// TIA Portal project "THELMA3_200224" (V15.1)

(* hardware
DEVICE "S71500/ET200MP station_1"  S7-1500 station
   slot 0: "Rail_0"  Rack  6ES7 590-1***0-0AA0
   slot 0: "PM 190W 120/230VAC"  PM 190W 120/230VAC  6EP1333-4BA00
   slot 1: "THELMA3"  CPU 1515-2 PN  6ES7 515-2AM01-0AB0  V2.6
      slot 3: "CPU display_1"  6ES7591-1BA00-0AA0
   slot 2: "DI 16x24VDC HF_1"  DI 16x24VDC HF  6ES7 521-1BH00-0AB0  V2.2
   slot 3: "DQ 16x24VDC/0.5A HF_1"  DQ 16x24VDC/0.5A HF  6ES7 522-1BH01-0AB0  V1.1
   slot 4: "DQ 16x24VDC/0.5A HF_2"  DQ 16x24VDC/0.5A HF  6ES7 522-1BH01-0AB0  V1.1
DEVICE "GSD device_1"  GSD.Device.PN
   slot 0: "Rack"  Rack  V1.0
   slot 0: "ucm8-bag-thelma3"  DataMan 260  DMR-260#-#0  5.5.0
      slot 0: "DataMan 260"  DataMan 260
      slot 1: "Interface"  Interface
         slot 1: "Port 1"  Port 1
   slot 1: "Acquisition Control_1"  Acquisition Control
      slot 0: "Acquisition Control"  Acquisition Control
   slot 2: "Acquisition Status_1"  Acquisition Status
      slot 0: "Acquisition Status"  Acquisition Status
   slot 3: "Results Control_1"  Results Control
      slot 0: "Results Control"  Results Control
   slot 4: "Results Status_1"  Results Status
      slot 0: "Results Status"  Results Status
   slot 5: "Soft Event Control_1"  Soft Event Control
      slot 0: "Soft Event Control"  Soft Event Control
   slot 6: "User Data - 64 bytes_1"  User Data - 64 bytes
      slot 0: "User Data - 64 bytes"  User Data - 64 bytes
   slot 7: "Result Data - 64 bytes_1"  Result Data - 64 bytes
      slot 0: "Result Data - 64 bytes"  Result Data - 64 bytes
DEVICE "GSD device_2"  GSD.Device.PN
   slot 0: "Rack"  Rack  V1.0
   slot 0: "ucm8-box-thelma3"  DataMan 260  DMR-260#-#0  5.5.0
      slot 0: "DataMan 260"  DataMan 260
      slot 1: "Interface"  Interface
         slot 1: "Port 1"  Port 1
   slot 1: "Acquisition Control_1"  Acquisition Control
      slot 0: "Acquisition Control"  Acquisition Control
   slot 2: "Acquisition Status_1"  Acquisition Status
      slot 0: "Acquisition Status"  Acquisition Status
   slot 3: "Results Control_1"  Results Control
      slot 0: "Results Control"  Results Control
   slot 4: "Results Status_1"  Results Status
      slot 0: "Results Status"  Results Status
   slot 5: "Soft Event Control_1"  Soft Event Control
      slot 0: "Soft Event Control"  Soft Event Control
   slot 6: "User Data - 128 bytes_1"  User Data - 128 bytes
      slot 0: "User Data - 128 bytes"  User Data - 128 bytes
   slot 7: "Result Data - 128 bytes_1"  Result Data - 128 bytes
      slot 0: "Result Data - 128 bytes"  Result Data - 128 bytes
DEVICE "HMI_THELMA3"  TP700 Comfort
   slot 0: "HMI_THELMA3"  TP700 Comfort  6AV2 124-0GC01-0AX0  15.1.0.0
   slot 1: "HMI_RT_2"  TP700 Comfort  6AV2 124-0GC01-0AX0  15.1.0.0
   slot 5: "HMI_THELMA3.1"  PROFINET Interface  15.0.1.0
      slot 1: "PROFINET Interface_1"  PROFINET Interface
         slot 1: "Port_1"  Port
         slot 2: "Port_2"  Port
   slot 7: "HMI_THELMA3._CP_1"  MPI/DP Interface  15.0.1.0
*)

// ===== PLC "THELMA3"  CPU 1515-2 PN =====

VAR_GLOBAL   // PLC tag table "Default tag table"
   "TrigerSensor" AT %I10.7 : Bool;
   "x_BypassPlainCheck" AT %M500.0 : Bool;
   "x_Arikel1" AT %M500.1 : Bool;
   "x_Artikel2" AT %M500.2 : Bool;
   "x_Artikel3" AT %M500.3 : Bool;
   "x_Artikel4" AT %M500.4 : Bool;
   "x_Simulacia_NoveData" AT %M505.0 : Bool;
   "x_Simulacia_Error" AT %M505.6 : Bool;
   "Kamera_odpojena" AT %M18.0 : Bool;
   "ArticleChangingBag" AT %M10.0 : Bool;
   "ArticleChangingBox" AT %M10.1 : Bool;
   "Reader2_Trigger_DelayTime" AT %MD68 : Time;
   "CON_HF_CommandTrigBatch" AT %M120.0 : Bool;
   "CON_HF_CommandTrig" AT %M120.1 : Bool;
   "CON_HF_CommandTrigBatchCon" AT %M120.2 : Bool;
   "CON_HF_CommandTrigAgainBatch" AT %M120.6 : Bool;
   "CON_HF_CommandTrigAgain" AT %M120.7 : Bool;
   "FirstScan" AT %M1.0 : Bool;
   "DiagStatusUpdate" AT %M1.1 : Bool;
   "TimeSynchPeriod" AT %MD64 : Time;
   "AlarmCheckPeriod" AT %MD60 : Time;
   "FaultByte1" AT %MB100 : Byte;
   "FaultByte2" AT %MB101 : Byte;
   "DelayTimeReader" AT %MD13 : Time;
   "CON_PrinterSelection" AT %M8.0 : Bool;
   "TRP_ErrorIP" AT %M105.0 : Bool;
   "TRP_CommError" AT %M105.1 : Bool;
   "TRP_HF_CommandTrig" AT %M121.1 : Bool;
   "TRP_ConnectHMI" AT %M121.4 : Bool;
   "TRP_HF_CommandTrigAgain" AT %M121.7 : Bool;
   "TRP_Inverse" AT %M140.0 : Bool;
   "TRP_Label" AT %M140.1 : Bool;
   "FaultByte3" AT %MB102 : Byte;
   "ResetFaults(1)" AT %M8.1 : Bool;
   "ResetCounters" AT %M8.2 : Bool;
   "CON_PrinterConnection" AT %M8.3 : Bool;
   "CON_ConnectHMI" AT %M120.4 : Bool;
   "System_Byte" AT %MB1 : Byte;
   "AlwaysTRUE" AT %M1.2 : Bool;
   "AlwaysFALSE" AT %M1.3 : Bool;
   "ResetResultAck" AT %M1500.0 : Bool;
   "LightYellowBag" AT %M50.0 : Bool;
   "LightYellowBox" AT %M51.0 : Bool;
   "LightRedBox" AT %M51.1 : Bool;
   "LightRedBag" AT %M50.1 : Bool;
   "LightGreenBox" AT %M51.2 : Bool;
   "LightGreenBag" AT %M50.2 : Bool;
   "NoReadCamBox" AT %M18.6 : Bool;   // IF NoRead <3 and Red light is off
   "Read_BOX_EM" AT %M52.0 : Bool;
   "Read_BOX_Enigma" AT %M52.1 : Bool;
   "Read_BOX_Mirai" AT %M52.2 : Bool;
   "SkuskaKroky" AT %MW1502 : Int;
   "PlainRedSignal" AT %M49.0 : Bool;
   "MIRAI_NoRead_A" AT %M107.0 : Bool;
   "MIRAI_MisMatch_A" AT %M107.1 : Bool;
   "LightRedMirai" AT %M51.3 : Bool;
   "FindRecipe" AT %M18.1 : Bool;   // bit pre automaticky vyber receptu
   "DataChange" AT %M18.2 : Bool;
   "TlacMDR" AT %M25.0 : Bool;
   "StatusCameraBag" AT %M18.4 : Bool;
   "StatusCameraBox" AT %M18.5 : Bool;
   "CamBagNoRead" AT %M21.0 : Bool;
   "NoReadCamBag" AT %M19.0 : Bool;   // IF NoRead <3 and Red light is off
END_VAR

VAR_GLOBAL   // PLC tag table "Bag"
   "Reader2_InspectionResults[0]" AT %IB400 : Byte;
   "Reader2_InspectionResults[1]" AT %IB401 : Byte;
   "Reader2_InspectionResults[2]" AT %IB402 : Byte;
   "Reader2_InspectionResults[3]" AT %IB403 : Byte;
   "Reader2_InspectionResults[4]" AT %IB404 : Byte;
   "Reader2_InspectionResults[5]" AT %IB405 : Byte;
   "Reader2_InspectionResults[6]" AT %IB406 : Byte;
   "Reader2_InspectionResults[7]" AT %IB407 : Byte;
   "Reader2_InspectionResults[8]" AT %IB408 : Byte;
   "Reader2_InspectionResults[9]" AT %IB409 : Byte;
   "Reader2_InspectionResults[10]" AT %IB410 : Byte;
   "Reader2_InspectionResults[11]" AT %IB411 : Byte;
   "Reader2_InspectionResults[12]" AT %IB412 : Byte;
   "Reader2_InspectionResults[13]" AT %IB413 : Byte;
   "Reader2_InspectionResults[14]" AT %IB414 : Byte;
   "Reader2_InspectionResults[15]" AT %IB415 : Byte;
   "Reader2_TriggerID" AT %IW121 : Word;
   "Reader2_Decoding" AT %I123.0 : Bool;
   "Reader2_DecodeComplete" AT %I123.1 : Bool;
   "Reader2_BufferOverrun" AT %I123.2 : Bool;
   "Reader2_ResultAvailable" AT %I123.3 : Bool;
   "Reader2_TrainCodeAck" AT %I124.0 : Bool;
   "Reader2_TrainMatchStrAck" AT %I124.1 : Bool;
   "Reader2_TrainFocusAck" AT %I124.2 : Bool;
   "Reader2_TrainBrightAck" AT %I124.3 : Bool;
   "Reader2_UnTrainAck" AT %I124.4 : Bool;
   "Reader2_ExecuteDmccAck" AT %I124.6 : Bool;
   "Reader2_SetMatchStringAck" AT %I124.7 : Bool;
   "Reader2_TriggerReady" AT %I120.0 : Bool;
   "Reader2_TriggerAck" AT %I120.1 : Bool;
   "Reader2_Acquiring" AT %I120.2 : Bool;
   "Reader2_MissedAquisition" AT %I120.3 : Bool;
   "Reader2_GeneralFault" AT %I123.7 : Bool;
   "Reader2_ResultID" AT %IW356 : Word;
   "Reader2_ResultCode" AT %IW358 : Word;
   "Reader2_ResultExtended" AT %IW360 : Word;
   "Reader2_Resultlength" AT %IW362 : Word;
   "Reader2_UserData[0]" AT %QB392 : Byte;
   "Reader2_UserData[1]" AT %QB393 : Byte;
   "Reader2_UserData[2]" AT %QB394 : Byte;
   "Reader2_UserData[3]" AT %QB395 : Byte;
   "Reader2_UserData[4]" AT %QB396 : Byte;
   "Reader2_UserData[5]" AT %QB397 : Byte;
   "Reader2_UserData[6]" AT %QB398 : Byte;
   "Reader2_UserData[7]" AT %QB399 : Byte;
   "Reader2_UserData[8]" AT %QB400 : Byte;
   "Reader2_UserData[9]" AT %QB401 : Byte;
   "Reader2_UserData[10]" AT %QB402 : Byte;
   "Reader2_UserData[11]" AT %QB403 : Byte;
   "Reader2_UserData[12]" AT %QB404 : Byte;
   "Reader2_UserData[13]" AT %QB405 : Byte;
   "Reader2_UserData[14]" AT %QB406 : Byte;
   "Reader2_UserData[15]" AT %QB407 : Byte;
   "Reader2_TriggerEnable" AT %Q120.0 : Bool;
   "Reader2_Trigger" AT %Q120.1 : Bool;
   "Reader2_BufferEnable" AT %Q121.0 : Bool;
   "Reader2_ResultsAck" AT %Q121.1 : Bool;
   "Reader2_TrainCode" AT %Q122.0 : Bool;
   "Reader2_TrainMatchString" AT %Q122.1 : Bool;
   "Reader2_TrainFocus" AT %Q122.2 : Bool;
   "Reader2_TrainBrightness" AT %Q122.3 : Bool;
   "Reader2_UnTrain" AT %Q122.4 : Bool;
   "Reader2_ExecuteDmcc" AT %Q122.6 : Bool;
   "Reader2_SetMatchString" AT %Q122.7 : Bool;
   "Reader2_UserDataOption" AT %QW388 : Word;
   "Reader2_UserDataLength" AT %QW390 : Word;
   "Reader2_UserData[16]" AT %QB408 : Byte;
   "Reader2_UserData[17]" AT %QB409 : Byte;
   "Reader2_UserData[18]" AT %QB410 : Byte;
   "Reader2_UserData[19]" AT %QB411 : Byte;
   "Reader2_UserData[20]" AT %QB412 : Byte;
   "Reader2_UserData[21]" AT %QB413 : Byte;
   "Reader2_UserData[22]" AT %QB414 : Byte;
   "Reader2_UserData[23]" AT %QB415 : Byte;
   "Reader2_UserData[24]" AT %QB416 : Byte;
   "Reader2_UserData[25]" AT %QB417 : Byte;
   "Reader2_UserData[26]" AT %QB418 : Byte;
   "Reader2_UserData[27]" AT %QB419 : Byte;
   "Reader2_UserData[28]" AT %QB420 : Byte;
   "Reader2_UserData[29]" AT %QB421 : Byte;
   "Reader2_UserData[30]" AT %QB422 : Byte;
   "Reader2_UserData[31]" AT %QB423 : Byte;
   "Reader2_UserData[32]" AT %QB424 : Byte;
   "Reader2_UserData[33]" AT %QB425 : Byte;
   "Reader2_UserData[34]" AT %QB426 : Byte;
   "Reader2_UserData[35]" AT %QB427 : Byte;
   "Reader2_UserData[36]" AT %QB428 : Byte;
   "Reader2_UserData[37]" AT %QB429 : Byte;
   "Reader2_UserData[38]" AT %QB430 : Byte;
   "Reader2_UserData[39]" AT %QB431 : Byte;
   "Reader2_UserData[40]" AT %QB432 : Byte;
   "LightYellowMirai" AT %M51.4 : Bool;
END_VAR

VAR_GLOBAL   // PLC tag table "Box"
   "Reader1_TriggerReady" AT %I110.0 : Bool;
   "Reader1_TriggerAck" AT %I110.1 : Bool;
   "Reader1_Acquiring" AT %I110.2 : Bool;
   "Reader1_MissedAcq" AT %I110.3 : Bool;
   "Reader1_TriggerID" AT %IW111 : Word;
   "Reader1_Decoding" AT %I113.0 : Bool;
   "Reader1_Decode Complete" AT %I113.1 : Bool;
   "Reader1_Results Buffer Overrun" AT %I113.2 : Bool;
   "Reader1_Results Available" AT %I113.3 : Bool;
   "Reader1_General Fault" AT %I113.7 : Bool;
   "Reader1_Train Code Ack" AT %I114.0 : Bool;
   "Reader1_Train Match String Ack" AT %I114.1 : Bool;
   "Reader1_Train Focus Ack" AT %I114.2 : Bool;
   "Reader1_Train Brightness Ack" AT %I114.3 : Bool;
   "Reader1_Untrain Ack" AT %I114.4 : Bool;
   "Reader1_Execute DMCC Ack" AT %I114.6 : Bool;
   "Reader1_Set Match String Ack" AT %I114.7 : Bool;
   "Reader1_ResultID" AT %IW256 : Word;
   "Reader1_Result Code" AT %IW258 : Word;
   "Reader1_Result Extended" AT %IW260 : Word;
   "Reader1_Result Length" AT %IW262 : Int;
   "Reader1_InspectionResults[0]" AT %IB264 : Byte;
   "Reader1_InspectionResults[1]" AT %IB265 : Byte;
   "Reader1_InspectionResults[2]" AT %IB266 : Byte;
   "Reader1_InspectionResults[3]" AT %IB267 : Byte;
   "Reader1_InspectionResults[4]" AT %IB268 : Byte;
   "Reader1_InspectionResults[5]" AT %IB269 : Byte;
   "Reader1_InspectionResults[6]" AT %IB270 : Byte;
   "Reader1_InspectionResults[7]" AT %IB271 : Byte;
   "Reader1_InspectionResults[8]" AT %IB272 : Byte;
   "Reader1_InspectionResults[9]" AT %IB273 : Byte;
   "Reader1_InspectionResults[10]" AT %IB274 : Byte;
   "Reader1_InspectionResults[11]" AT %IB275 : Byte;
   "Reader1_InspectionResults[12]" AT %IB276 : Byte;
   "Reader1_InspectionResults[13]" AT %IB277 : Byte;
   "Reader1_InspectionResults[14]" AT %IB278 : Byte;
   "Reader1_InspectionResults[15]" AT %IB279 : Byte;
   "Reader1_InspectionResults[16]" AT %IB280 : Byte;
   "Reader1_InspectionResults[17]" AT %IB281 : Byte;
   "Reader1_InspectionResults[18]" AT %IB282 : Byte;
   "Reader1_InspectionResults[19]" AT %IB283 : Byte;
   "Reader1_InspectionResults[20]" AT %IB284 : Byte;
   "Reader1_InspectionResults[21]" AT %IB285 : Byte;
   "Reader1_InspectionResults[22]" AT %IB286 : Byte;
   "Reader1_InspectionResults[23]" AT %IB287 : Byte;
   "Reader1_InspectionResults[24]" AT %IB288 : Byte;
   "Reader1_InspectionResults[25]" AT %IB289 : Byte;
   "Reader1_InspectionResults[26]" AT %IB290 : Byte;
   "Reader1_InspectionResults[27]" AT %IB291 : Byte;
   "Reader1_InspectionResults[28]" AT %IB292 : Byte;
   "Reader1_InspectionResults[29]" AT %IB293 : Byte;
   "Reader1_InspectionResults[30]" AT %IB294 : Byte;
   "Reader1_InspectionResults[31]" AT %IB295 : Byte;
   "Reader1_InspectionResults[32]" AT %IB296 : Byte;
   "Reader1_InspectionResults[33]" AT %IB297 : Byte;
   "Reader1_InspectionResults[34]" AT %IB298 : Byte;
   "Reader1_InspectionResults[35]" AT %IB299 : Byte;
   "Reader1_InspectionResults[36]" AT %IB300 : Byte;
   "Reader1_InspectionResults[37]" AT %IB301 : Byte;
   "Reader1_InspectionResults[38]" AT %IB302 : Byte;
   "Reader1_InspectionResults[39]" AT %IB303 : Byte;
   "Reader1_InspectionResults[40]" AT %IB304 : Byte;
   "Reader1_InspectionResults[41]" AT %IB305 : Byte;
   "Reader1_InspectionResults[42]" AT %IB306 : Byte;
   "Reader1_InspectionResults[43]" AT %IB307 : Byte;
   "Reader1_InspectionResults[44]" AT %IB308 : Byte;
   "Reader1_InspectionResults[45]" AT %IB309 : Byte;
   "Reader1_InspectionResults[46]" AT %IB310 : Byte;
   "Reader1_InspectionResults[47]" AT %IB311 : Byte;
   "Reader1_InspectionResults[48]" AT %IB312 : Byte;
   "Reader1_InspectionResults[49]" AT %IB313 : Byte;
   "Reader1_InspectionResults[50]" AT %IB314 : Byte;
   "Reader1_InspectionResults[51]" AT %IB315 : Byte;
   "Reader1_InspectionResults[52]" AT %IB316 : Byte;
   "Reader1_InspectionResults[53]" AT %IB317 : Byte;
   "Reader1_InspectionResults[54]" AT %IB318 : Byte;
   "Reader1_InspectionResults[55]" AT %IB319 : Byte;
   "Reader1_InspectionResults[56]" AT %IB320 : Byte;
   "Reader1_InspectionResults[57]" AT %IB321 : Byte;
   "Reader1_InspectionResults[58]" AT %IB322 : Byte;
   "Reader1_InspectionResults[59]" AT %IB323 : Byte;
   "Reader1_InspectionResults[60]" AT %IB324 : Byte;
   "Reader1_InspectionResults[61]" AT %IB325 : Byte;
   "Reader1_InspectionResults[62]" AT %IB326 : Byte;
   "Reader1_InspectionResults[63]" AT %IB327 : Byte;
   "Reader1_InspectionResults[64]" AT %IB328 : Byte;
   "Reader1_InspectionResults[65]" AT %IB329 : Byte;
   "Reader1_InspectionResults[66]" AT %IB330 : Byte;
   "Reader1_InspectionResults[67]" AT %IB331 : Byte;
   "Reader1_InspectionResults[68]" AT %IB332 : Byte;
   "Reader1_InspectionResults[69]" AT %IB333 : Byte;
   "Reader1_InspectionResults[70]" AT %IB334 : Byte;
   "Reader1_InspectionResults[71]" AT %IB335 : Byte;
   "Reader1_InspectionResults[72]" AT %IB336 : Byte;
   "Reader1_InspectionResults[73]" AT %IB337 : Byte;
   "Reader1_InspectionResults[74]" AT %IB338 : Byte;
   "Reader1_InspectionResults[75]" AT %IB339 : Byte;
   "Reader1_InspectionResults[76]" AT %IB340 : Byte;
   "Reader1_InspectionResults[77]" AT %IB341 : Byte;
   "Reader1_InspectionResults[78]" AT %IB342 : Byte;
   "Reader1_InspectionResults[79]" AT %IB343 : Byte;
   "Reader1_InspectionResults[80]" AT %IB344 : Byte;
   "Reader1_InspectionResults[81]" AT %IB345 : Byte;
   "Reader1_InspectionResults[82]" AT %IB346 : Byte;
   "Reader1_InspectionResults[83]" AT %IB347 : Byte;
   "Reader1_InspectionResults[84]" AT %IB348 : Byte;
   "Reader1_InspectionResults[85]" AT %IB349 : Byte;
   "Reader1_InspectionResults[86]" AT %IB350 : Byte;
   "Reader1_InspectionResults[87]" AT %IB351 : Byte;
   "Reader1_InspectionResults[88]" AT %IB352 : Byte;
   "Reader1_InspectionResults[89]" AT %IB353 : Byte;
   "Reader1_InspectionResults[90]" AT %IB354 : Byte;
   "Reader1_InspectionResults[91]" AT %IB355 : Byte;
   "Reader1_InspectionResults[92]" AT %IB356 : Byte;
   "Reader1_InspectionResults[93]" AT %IB357 : Byte;
   "Reader1_InspectionResults[94]" AT %IB358 : Byte;
   "Reader1_InspectionResults[95]" AT %IB359 : Byte;
   "Reader1_InspectionResults[96]" AT %IB360 : Byte;
   "Reader1_InspectionResults[97]" AT %IB361 : Byte;
   "Reader1_InspectionResults[98]" AT %IB362 : Byte;
   "Reader1_InspectionResults[99]" AT %IB363 : Byte;
   "Reader1_InspectionResults[100]" AT %IB364 : Byte;
   "Reader1_InspectionResults[101]" AT %IB365 : Byte;
   "Reader1_InspectionResults[102]" AT %IB366 : Byte;
   "Reader1_InspectionResults[103]" AT %IB367 : Byte;
   "Reader1_InspectionResults[104]" AT %IB368 : Byte;
   "Reader1_InspectionResults[105]" AT %IB369 : Byte;
   "Reader1_InspectionResults[106]" AT %IB370 : Byte;
   "Reader1_InspectionResults[107]" AT %IB371 : Byte;
   "Reader1_InspectionResults[108]" AT %IB372 : Byte;
   "Reader1_InspectionResults[109]" AT %IB373 : Byte;
   "Reader1_InspectionResults[110]" AT %IB374 : Byte;
   "Reader1_InspectionResults[111]" AT %IB375 : Byte;
   "Reader1_InspectionResults[112]" AT %IB376 : Byte;
   "Reader1_InspectionResults[113]" AT %IB377 : Byte;
   "Reader1_InspectionResults[114]" AT %IB378 : Byte;
   "Reader1_InspectionResults[115]" AT %IB379 : Byte;
   "Reader1_InspectionResults[116]" AT %IB380 : Byte;
   "Reader1_InspectionResults[117]" AT %IB381 : Byte;
   "Reader1_InspectionResults[118]" AT %IB382 : Byte;
   "Reader1_InspectionResults[119]" AT %IB383 : Byte;
   "Reader1_InspectionResults[120]" AT %IB384 : Byte;
   "Reader1_InspectionResults[121]" AT %IB385 : Byte;
   "Reader1_InspectionResults[122]" AT %IB386 : Byte;
   "Reader1_InspectionResults[123]" AT %IB387 : Byte;
   "Reader1_InspectionResults[124]" AT %IB388 : Byte;
   "Reader1_InspectionResults[125]" AT %IB389 : Byte;
   "Reader1_InspectionResults[126]" AT %IB390 : Byte;
   "Reader1_InspectionResults[127]" AT %IB391 : Byte;
   "Reader1_TriggerEnable" AT %Q110.0 : Bool;
   "Reader1_Trigger" AT %Q110.1 : Bool;
   "Reader1_BufferResultsEnable" AT %Q111.0 : Bool;
   "Reader1_ResultsAck" AT %Q111.1 : Bool;
   "Reader1_Train Code" AT %Q112.0 : Bool;
   "Reader1_Train Match String" AT %Q112.1 : Bool;
   "Reader1_Train Focus" AT %Q112.2 : Bool;
   "Reader1_Train Brightness" AT %Q112.3 : Bool;
   "Reader1_Untrain" AT %Q112.4 : Bool;
   "Reader1_Execute DMCC" AT %Q112.6 : Bool;
   "Reader1_Set Match String" AT %Q112.7 : Bool;
   "Reader1_UserData Option" AT %QW256 : Word;
   "Reader1_UserData Length" AT %QW258 : Word;
   "Reader1_UserData[0]" AT %QB260 : Byte;
   "Reader1_UserData[1]" AT %QB261 : Byte;
   "Reader1_UserData[2]" AT %QB262 : Byte;
   "Reader1_UserData[3]" AT %QB263 : Byte;
   "Reader1_UserData[4]" AT %QB264 : Byte;
   "Reader1_UserData[5]" AT %QB265 : Byte;
   "Reader1_UserData[6]" AT %QB266 : Byte;
   "Reader1_UserData[7]" AT %QB267 : Byte;
   "Reader1_UserData[8]" AT %QB268 : Byte;
   "Reader1_UserData[9]" AT %QB269 : Byte;
   "Reader1_UserData[10]" AT %QB270 : Byte;
   "Reader1_UserData[11]" AT %QB271 : Byte;
   "Reader1_UserData[12]" AT %QB272 : Byte;
   "Reader1_UserData[13]" AT %QB273 : Byte;
   "Reader1_UserData[14]" AT %QB274 : Byte;
   "Reader1_UserData[15]" AT %QB275 : Byte;
   "Reader1_UserData[16]" AT %QB276 : Byte;
   "Reader1_UserData[17]" AT %QB277 : Byte;
   "Reader1_UserData[18]" AT %QB278 : Byte;
   "Reader1_UserData[19]" AT %QB279 : Byte;
   "Reader1_UserData[20]" AT %QB280 : Byte;
   "Reader1_UserData[21]" AT %QB281 : Byte;
   "Reader1_UserData[22]" AT %QB282 : Byte;
   "Reader1_UserData[23]" AT %QB283 : Byte;
   "Reader1_UserData[24]" AT %QB284 : Byte;
   "Reader1_UserData[25]" AT %QB285 : Byte;
   "Reader1_UserData[26]" AT %QB286 : Byte;
   "Reader1_UserData[27]" AT %QB287 : Byte;
   "Reader1_UserData[28]" AT %QB288 : Byte;
   "Reader1_UserData[29]" AT %QB289 : Byte;
   "Reader1_UserData[30]" AT %QB290 : Byte;
   "Reader1_UserData[31]" AT %QB291 : Byte;
   "Reader1_UserData[32]" AT %QB292 : Byte;
   "Reader1_UserData[33]" AT %QB293 : Byte;
   "Reader1_UserData[34]" AT %QB294 : Byte;
   "Reader1_UserData[35]" AT %QB295 : Byte;
   "Reader1_UserData[36]" AT %QB296 : Byte;
   "Reader1_UserData[37]" AT %QB297 : Byte;
   "Reader1_UserData[38]" AT %QB298 : Byte;
   "Reader1_UserData[39]" AT %QB299 : Byte;
   "Reader1_UserData[40]" AT %QB300 : Byte;
   "Reader1_UserData[41]" AT %QB301 : Byte;
   "Reader1_UserData[42]" AT %QB302 : Byte;
   "Reader1_UserData[43]" AT %QB303 : Byte;
   "Reader1_UserData[44]" AT %QB304 : Byte;
   "Reader1_UserData[45]" AT %QB305 : Byte;
   "Reader1_UserData[46]" AT %QB306 : Byte;
   "Reader1_UserData[47]" AT %QB307 : Byte;
   "Reader1_UserData[48]" AT %QB308 : Byte;
   "Reader1_UserData[49]" AT %QB309 : Byte;
   "Reader1_UserData[50]" AT %QB310 : Byte;
   "Reader1_UserData[51]" AT %QB311 : Byte;
   "Reader1_UserData[52]" AT %QB312 : Byte;
   "Reader1_UserData[53]" AT %QB313 : Byte;
   "Reader1_UserData[54]" AT %QB314 : Byte;
   "Reader1_UserData[55]" AT %QB315 : Byte;
   "Reader1_UserData[56]" AT %QB316 : Byte;
   "Reader1_UserData[57]" AT %QB317 : Byte;
   "Reader1_UserData[58]" AT %QB318 : Byte;
   "Reader1_UserData[59]" AT %QB319 : Byte;
   "Reader1_UserData[60]" AT %QB320 : Byte;
   "Reader1_UserData[61]" AT %QB321 : Byte;
   "Reader1_UserData[62]" AT %QB322 : Byte;
   "Reader1_UserData[63]" AT %QB323 : Byte;
   "Reader1_UserData[64]" AT %QB324 : Byte;
   "Reader1_UserData[65]" AT %QB325 : Byte;
   "Reader1_UserData[66]" AT %QB326 : Byte;
   "Reader1_UserData[67]" AT %QB327 : Byte;
   "Reader1_UserData[68]" AT %QB328 : Byte;
   "Reader1_UserData[69]" AT %QB329 : Byte;
   "Reader1_UserData[70]" AT %QB330 : Byte;
   "Reader1_UserData[71]" AT %QB331 : Byte;
   "Reader1_UserData[72]" AT %QB332 : Byte;
   "Reader1_UserData[73]" AT %QB333 : Byte;
   "Reader1_UserData[74]" AT %QB334 : Byte;
   "Reader1_UserData[75]" AT %QB335 : Byte;
   "Reader1_UserData[76]" AT %QB336 : Byte;
   "Reader1_UserData[77]" AT %QB337 : Byte;
   "Reader1_UserData[78]" AT %QB338 : Byte;
   "Reader1_UserData[79]" AT %QB339 : Byte;
   "Reader1_UserData[80]" AT %QB340 : Byte;
   "Reader1_UserData[81]" AT %QB341 : Byte;
   "Reader1_UserData[82]" AT %QB342 : Byte;
   "Reader1_UserData[83]" AT %QB343 : Byte;
   "Reader1_UserData[84]" AT %QB344 : Byte;
   "Reader1_UserData[85]" AT %QB345 : Byte;
   "Reader1_UserData[86]" AT %QB346 : Byte;
   "Reader1_UserData[87]" AT %QB347 : Byte;
   "Reader1_UserData[88]" AT %QB348 : Byte;
   "Reader1_UserData[89]" AT %QB349 : Byte;
   "Reader1_UserData[90]" AT %QB350 : Byte;
   "Reader1_UserData[91]" AT %QB351 : Byte;
   "Reader1_UserData[92]" AT %QB352 : Byte;
   "Reader1_UserData[93]" AT %QB353 : Byte;
   "Reader1_UserData[94]" AT %QB354 : Byte;
   "Reader1_UserData[95]" AT %QB355 : Byte;
   "Reader1_UserData[96]" AT %QB356 : Byte;
   "Reader1_UserData[97]" AT %QB357 : Byte;
   "Reader1_UserData[98]" AT %QB358 : Byte;
   "Reader1_UserData[99]" AT %QB359 : Byte;
   "Reader1_UserData[100]" AT %QB360 : Byte;
   "Reader1_UserData[101]" AT %QB361 : Byte;
   "Reader1_UserData[102]" AT %QB362 : Byte;
   "Reader1_UserData[103]" AT %QB363 : Byte;
   "Reader1_UserData[104]" AT %QB364 : Byte;
   "Reader1_UserData[105]" AT %QB365 : Byte;
   "Reader1_UserData[106]" AT %QB366 : Byte;
   "Reader1_UserData[107]" AT %QB367 : Byte;
   "Reader1_UserData[108]" AT %QB368 : Byte;
   "Reader1_UserData[109]" AT %QB369 : Byte;
   "Reader1_UserData[110]" AT %QB370 : Byte;
   "Reader1_UserData[111]" AT %QB371 : Byte;
   "Reader1_UserData[112]" AT %QB372 : Byte;
   "Reader1_UserData[113]" AT %QB373 : Byte;
   "Reader1_UserData[114]" AT %QB374 : Byte;
   "Reader1_UserData[115]" AT %QB375 : Byte;
   "Reader1_UserData[116]" AT %QB376 : Byte;
   "Reader1_UserData[117]" AT %QB377 : Byte;
   "Reader1_UserData[118]" AT %QB378 : Byte;
   "Reader1_UserData[119]" AT %QB379 : Byte;
   "Reader1_UserData[120]" AT %QB380 : Byte;
   "Reader1_UserData[121]" AT %QB381 : Byte;
   "Reader1_UserData[122]" AT %QB382 : Byte;
   "Reader1_UserData[123]" AT %QB383 : Byte;
   "Reader1_UserData[124]" AT %QB384 : Byte;
   "Reader1_UserData[125]" AT %QB385 : Byte;
   "Reader1_UserData[126]" AT %QB386 : Byte;
   "Reader1_UserData[127]" AT %QB387 : Byte;
END_VAR

VAR_GLOBAL   // PLC tag table "In"
   "Lable_tlac_istic" AT %I10.0 : Bool;
   "DI_napajanie_24V" AT %I10.1 : Bool;
   "Ventilator_napajanie" AT %I10.2 : Bool;
   "Cam_BAG_trigger" AT %I10.4 : Bool;
   "Cam_BAG_kod_Read" AT %I10.5 : Bool;
   "Cam_BAG_kod_NoRead" AT %I10.6 : Bool;
   "Cam_BOX_trigger" AT %I11.0 : Bool;
   "Cam_BOX_kod_Read" AT %I11.1 : Bool;
   "Cam_BOX_kod_NoRead" AT %I11.2 : Bool;
END_VAR

VAR_GLOBAL   // PLC tag table "Out"
   "BAG_MisMatch" AT %Q10.0 : Bool;
   "BAG_NoValidated" AT %Q10.1 : Bool;
   "BAG_NoRead" AT %Q10.2 : Bool;
   "BAG_CodeNotPressent" AT %Q10.3 : Bool;
   "BAG_CameraNotReady" AT %Q10.4 : Bool;
   "BAG_TriggerNotReady" AT %Q10.5 : Bool;
   "BOX_MisMatch" AT %Q10.6 : Bool;
   "BOX_NoValidated" AT %Q10.7 : Bool;
   "BOX_NoRead" AT %Q11.0 : Bool;
   "BOX_CodeNotPresent" AT %Q11.1 : Bool;
   "BOX_CameraNotReady" AT %Q11.2 : Bool;
   "BOX_TriggerNotReady" AT %Q11.3 : Bool;
   "LightGreen" AT %Q11.4 : Bool;
   "LightYellow" AT %Q11.5 : Bool;
   "LightRed" AT %Q11.6 : Bool;
   "MIRAI_MisMatch" AT %Q14.0 : Bool;
   "MIRAI_NoRead" AT %Q14.1 : Bool;
   "MIRAI_FaultLablePrinter" AT %Q14.2 : Bool;
   "MIRAI_AlarmLablePrinter" AT %Q14.3 : Bool;
   "MIRAI_FaultVideoJet" AT %Q14.4 : Bool;
   "MIRAI_AlarmVideoJet" AT %Q14.5 : Bool;
   "MIRAI_OPC_ERROR" AT %Q14.6 : Bool;
END_VAR

VAR_GLOBAL CONSTANT   // PLC tag table "Default tag table_1"
   "None(1)" : Pip := 65535;
   "Automatic update(1)" : Pip := 0;
   "PIP 1(1)" : Pip := 1;
   "PIP 2(1)" : Pip := 2;
   "PIP 3(1)" : Pip := 3;
   "PIP 4(1)" : Pip := 4;
   "PIP 5(1)" : Pip := 5;
   "PIP 6(1)" : Pip := 6;
   "PIP 7(1)" : Pip := 7;
   "PIP 8(1)" : Pip := 8;
   "PIP 9(1)" : Pip := 9;
   "PIP 10(1)" : Pip := 10;
   "PIP 11(1)" : Pip := 11;
   "PIP 12(1)" : Pip := 12;
   "PIP 13(1)" : Pip := 13;
   "PIP 14(1)" : Pip := 14;
   "PIP 15(1)" : Pip := 15;
   "PIP 16(1)" : Pip := 16;
   "PIP 17(1)" : Pip := 17;
   "PIP 18(1)" : Pip := 18;
   "PIP 19(1)" : Pip := 19;
   "PIP 20(1)" : Pip := 20;
   "PIP 21(1)" : Pip := 21;
   "PIP 22(1)" : Pip := 22;
   "PIP 23(1)" : Pip := 23;
   "PIP 24(1)" : Pip := 24;
   "PIP 25(1)" : Pip := 25;
   "PIP 26(1)" : Pip := 26;
   "PIP 27(1)" : Pip := 27;
   "PIP 28(1)" : Pip := 28;
   "PIP 29(1)" : Pip := 29;
   "PIP 30(1)" : Pip := 30;
   "PIP 31(1)" : Pip := 31;
   "PIP OB Servo(1)" : Pip := 32768;
   "Local~Exec(1)" : Hw_SubModule := 52;
   "Local(1)" : Hw_SubModule := 49;
   "Local~PROFINET_interface_1~Port_2(1)" : Hw_Interface := 66;
   "Local~DI_16x24VDC_HF_1(1)" : Hw_SubModule := 259;
   "Local~DQ_16x24VDC_0_5A_HF_1" : Hw_SubModule := 260;
   "Local~PROFINET_IO-System(1)" : Hw_IoSystem := 258;
   "ucm8-box-dm262~Proxy(1)" : Hw_SubModule := 266;
   "ucm8-box-dm262~IODevice(1)" : Hw_Device := 262;
   "ucm8-box-dm262~Interface(1)" : Hw_Interface := 268;
   "ucm8-box-dm262~Interface~Port_1(1)" : Hw_Interface := 270;
   "ucm8-box-dm262~Head(1)" : Hw_SubModule := 261;
   "ucm8-box-dm262~Acquisition_Control_1(1)" : Hw_SubModule := 263;
   "ucm8-box-dm262~Acquisition_Status_1(1)" : Hw_SubModule := 265;
   "ucm8-box-dm262~Results_Control_1(1)" : Hw_SubModule := 267;
   "ucm8-box-dm262~Results_Status_1(1)" : Hw_SubModule := 269;
   "ucm8-box-dm262~Soft_Event_Control_1(1)" : Hw_SubModule := 271;
   "ucm8-box-dm262~User_Data_-_64_bytes_1" : Hw_SubModule := 273;
   "ucm8-box-dm262~Result_Data_-_64_bytes_1" : Hw_SubModule := 275;
   "Local~PM_70W_120_230VAC" : Hw_SubModule := 257;
   "Local~Display(1)" : Hw_SubModule := 54;
   "Local~MC(1)" : Hw_SubModule := 51;
   "Local~PROFINET_interface_1(1)" : Hw_Interface := 64;
   "Local~PROFINET_interface_1~Port_1(1)" : Hw_Interface := 65;
   "Local~Common(1)" : Hw_SubModule := 50;
   "Local~Device(1)" : Hw_Device := 32;
   "Local~Configuration(1)" : Hw_SubModule := 33;
   "ucm8-bag-dm262~Proxy(1)" : Hw_SubModule := 276;
   "ucm8-bag-dm262~IODevice(1)" : Hw_Device := 272;
   "ucm8-bag-dm262~Interface(1)" : Hw_Interface := 277;
   "ucm8-bag-dm262~Interface~Port_1(1)" : Hw_Interface := 278;
   "ucm8-bag-dm262~Head(1)" : Hw_SubModule := 279;
   "ucm8-bag-dm262~Acquisition_Control_1(1)" : Hw_SubModule := 280;
   "ucm8-bag-dm262~Acquisition_Status_1(1)" : Hw_SubModule := 281;
   "ucm8-bag-dm262~Results_Control_1(1)" : Hw_SubModule := 282;
   "ucm8-bag-dm262~Results_Status_1(1)" : Hw_SubModule := 283;
   "ucm8-bag-dm262~Soft_Event_Control_1(1)" : Hw_SubModule := 284;
   "ucm8-bag-dm262~User_Data_-_64_bytes_1(1)" : Hw_SubModule := 285;
   "ucm8-bag-dm262~Result_Data_-_64_bytes_1(1)" : Hw_SubModule := 286;
   "OB_Startup" : OB_STARTUP := 100;
   "OB_RackStationFailure(1)" : OB_Any := 86;
   "OB_Main(1)" : OB_PCYCLE := 1;
END_VAR

VAR_GLOBAL   // PLC tag table "Common"
   "Clock_Byte" AT %MB255 : Byte;
   "Clock_10Hz" AT %M255.0 : Bool;
   "Clock_5Hz" AT %M255.1 : Bool;
   "Clock_2.5Hz" AT %M255.2 : Bool;
   "Clock_2Hz" AT %M255.3 : Bool;
   "Clock_1.25Hz" AT %M255.4 : Bool;
   "Clock_1Hz" AT %M255.5 : Bool;
   "Clock_0.625Hz" AT %M255.6 : Bool;
   "Clock_0.5Hz" AT %M255.7 : Bool;
END_VAR

VAR_GLOBAL   // PLC tag table "Faults"
   "Box_FltMisMatch" AT %M101.1 : Bool;
   "Box_FltNoRead" AT %M101.2 : Bool;
   "FltAccessIO" AT %M101.0 : Bool;
   "Box_FltTriggerWatchDog" AT %M101.3 : Bool;
   "Box_MsgNoRead" AT %M111.2 : Bool;
   "Bag_FltMisMatch" AT %M103.1 : Bool;
   "Bag_FltNoRead" AT %M103.2 : Bool;
   "Bag_FltTriggerWatchDog" AT %M103.3 : Bool;
   "Bag_MsgNoRead" AT %M112.2 : Bool;
   "FaultWord1" AT %MW100 : Word;
   "FaultWord2" AT %MW102 : Word;
   "FaultWord3" AT %MW104 : Word;
   "FaultWord4" AT %MW106 : Word;
   "FaultWord5" AT %MW108 : Word;
   "FaultWord6" AT %MW110 : Word;
   "FaultWord7" AT %MW112 : Word;
   "FaultWord8" AT %MW114 : Word;
   "BoxEnigmaDisable" AT %M101.4 : Bool;
   "BagEnigmaDisable" AT %M103.4 : Bool;
   "BagMaterialNumberNotValid" AT %M103.5 : Bool;
   "BoxMaterialNumberNotValid" AT %M101.5 : Bool;
   "CON_ErrorIP" AT %M100.0 : Bool;
   "Hw_Fault" AT %M110.5 : Bool;
   "PLAIN_ERROR" AT %M100.4 : Bool;
   "Lable_print_Istic" AT %M106.0 : Bool;
   "Napajanie_DI" AT %M106.1 : Bool;
   "Napajanie_ventilator" AT %M106.2 : Bool;
   "LiveBitError" AT %M100.5 : Bool;
   "NoNewData" AT %M100.6 : Bool;
   "BatchEndTimeWarning" AT %M102.0 : Bool;
   "BatchEndTimeError" AT %M102.1 : Bool;
   "FaultCamBag" AT %M111.0 : Bool;
   "FaultCamBox" AT %M111.1 : Bool;
   "Overheated" AT %M108.0 : Bool;
   "IO_BoardError" AT %M108.1 : Bool;
   "FileSystemError" AT %M108.2 : Bool;
   "MemoryError" AT %M108.3 : Bool;
   "ParameterError" AT %M108.4 : Bool;
   "NoInitError" AT %M108.5 : Bool;
   "NoAirPressure" AT %M108.6 : Bool;
   "PaperOut" AT %M108.7 : Bool;
   "RibbonOut" AT %M109.0 : Bool;
   "HeadLifted" AT %M109.1 : Bool;
   "PressStart" AT %M109.2 : Bool;
   "NoReturnSignal" AT %M109.3 : Bool;
   "ArmJammed" AT %M109.4 : Bool;
   "ArmNotHome" AT %M109.5 : Bool;
   "BarcodeError" AT %M109.6 : Bool;
   "LabelOnGrid" AT %M109.7 : Bool;
   "NoLabelOnGrid" AT %M114.0 : Bool;
   "CoverOpen" AT %M114.1 : Bool;
   "Pause" AT %M114.2 : Bool;
   "PaperLow" AT %M114.3 : Bool;
   "RibbonLow" AT %M114.4 : Bool;
   "BarcodeWarning" AT %M114.5 : Bool;
   "ApplyDelayTooShort" AT %M114.6 : Bool;
   "AcceptDateChange" AT %M114.7 : Bool;
   "MatchCodeError" AT %M115.0 : Bool;
   "BarcodeQuality" AT %M115.1 : Bool;
   "WaitingForTrig" AT %M115.2 : Bool;
   "TrigSensorError" AT %M115.3 : Bool;
   "PrinterSynchronization" AT %M115.4 : Bool;
   "SynchronizationTimeout" AT %M115.5 : Bool;
   "ProductToClose" AT %M115.6 : Bool;
   "SSCC_LimitReached" AT %M115.7 : Bool;
END_VAR

VAR_GLOBAL CONSTANT   // PLC tag table "LCom_Constants"
   "LCOM_NO_TIME_SYNC" : USInt := 0;
   "LCOM_TCP_CONNECTION" : USInt := 1;
   "LCOM_LCOM_CONNECTION" : USInt := 2;
   "LCOM_CYCLE_TIME_SYNC" : USInt := 1;
   "LCOM_TIME_OF_DAY_TIME_SYNC" : USInt := 2;
   "LCOM_STATUS_NO_CALL" : Word := 16#7000;
   "LCOM_STATUS_FIRST_CALL" : Word := 16#7001;
   "LCOM_STATUS_INTERMEDIATE_CALL" : Word := 16#7002;
   "LCOM_STATUS_CLIENT_TRY_CONNECT" : Word := 16#7003;
   "LCOM_STATUS_SERVER_PORT_OPEN" : Word := 16#7004;
   "LCOM_STATUS_TCP_CONNECTED" : Word := 16#7005;
   "LCOM_STATUS_LCOM_CONNECTED_V1" : Word := 16#7006;
   "LCOM_STATUS_LCOM_CONNECTED_V2" : Word := 16#7007;
   "LCOM_STATUS_DISCONNECTING" : Word := 16#7008;
   "LCOM_WARN_SEND_DATA_LENGTH" : Word := 16#7600;
   "LCOM_WARN_LIFE_SIGN_LIMITATION" : Word := 16#7610;
   "LCOM_WARN_SEND_CYCLE_LIMITATION" : Word := 16#7611;
   "LCOM_WARN_ACK_TIMEOUT_LIMITATION" : Word := 16#7612;
   "LCOM_WARN_SEND_CYCLE_EXPIRED" : Word := 16#7613;
   "LCOM_WARN_RECEIVE_BUFFER_LEN" : Word := 16#7614;
   "LCOM_WARN_NO_TIME_SYNC" : Word := 16#7615;
   "LCOM_ERR_COM_SERVICE" : Word := 16#8200;
   "LCOM_ERR_CONNECTION_ID" : Word := 16#8201;
   "LCOM_ERR_INTERFACE_ID" : Word := 16#8202;
   "LCOM_ERR_LOCAL_PORT" : Word := 16#8203;
   "LCOM_ERR_PARTNER_IP" : Word := 16#8204;
   "LCOM_ERR_TIME_SYNC_MODE" : Word := 16#8205;
   "LCOM_ERR_TIME_CYCLE_TIME" : Word := 16#8206;
   "LCOM_ERR_TIME_OF_DAY" : Word := 16#8207;
   "LCOM_ERR_SEND_DATA_TYPE" : Word := 16#8208;
   "LCOM_ERR_RECEIVE_DATA_TYPE" : Word := 16#8209;
   "LCOM_ERR_LIFE_SIGN_CYCLE" : Word := 16#8210;
   "LCOM_ERR_SEND_CYCLE_TIME" : Word := 16#8211;
   "LCOM_ERR_ACK_TIMEOUT" : Word := 16#8212;
   "LCOM_ERR_OPEN_CLIENT" : Word := 16#8600;
   "LCOM_ERR_OPEN_SERVER" : Word := 16#8601;
   "LCOM_ERR_SEND" : Word := 16#8602;
   "LCOM_ERR_RECEIVE" : Word := 16#8603;
   "LCOM_ERR_CLOSE_CONNECTION" : Word := 16#8604;
   "LCOM_ERR_LIFE_SIGN_EXPIRED" : Word := 16#8610;
   "LCOM_ERR_ACK_TIMEOUT_EXPIRED" : Word := 16#8611;
   "LCOM_ERR_ACK_MESSAGE_NUMBER" : Word := 16#8612;
   "LCOM_ERR_WRONG_LCOM_HEADER" : Word := 16#8613;
   "LCOM_ERR_WRONG_TELEGRAM_ID" : Word := 16#8614;
END_VAR

VAR_GLOBAL   // PLC tag table "Tag table_1"
   "CON_CommError" AT %M100.1 : Bool;
END_VAR

TYPE "UDT_Printer"
VERSION : 0.1
   STRUCT
      RemoteAddress : String;
      "Date" : String;
      "Time" : String;
      RData : Array[0..56] of Byte;
      RdataBatch : Array[0..56] of Byte;
      BatchOK : Bool;
      TimeOK : Bool;
      NoAlarm : Bool;
      LED_State : USInt;
      TimeDateError : Bool;
      OPC_Error : Bool;
      TCP_ComError : Bool;
      Inverse : Bool;
      Initialization : Bool;
      TCP_ComErrorBatch : Bool;
      ComErrorStatus : Byte;
      ComErrorStatusBatch : Byte;
   END_STRUCT;
END_TYPE

TYPE "UDT_LatestReadingBag"
VERSION : 0.1
   STRUCT
      ID : Int;
      Flags : Int;
      Length : Int;
      Value : Array[0..9] of Char;
   END_STRUCT;
END_TYPE

TYPE "UDT_CON_Comm"
VERSION : 0.1
   STRUCT
      Heartbeat : Bool;
      HeartbeatToPlain : Bool;
      NewMDR_Flag : String;
      NewArticleFlag : String;
      NewBatchNumber : String;
      NewArtBaseNumber : UDInt;
      NewMarketREG_Code : String;
      NewBatchEndTime : String;
      NewBBD : String;
      ActualBatchNumber : String;
      ActualArtBaseNumber : String;
      ActualMarketRegCode : String;
      ActualBBD : String;
      BatchStatus : Byte;
   END_STRUCT;
END_TYPE

TYPE "UDT_Reader"
VERSION : 0.1
   STRUCT
      ResetFaults : Bool;
      ResetCounters : Bool;
      MisMatchFault : Bool;
      NoReadFault : Bool;
      MisTriggerFault : Bool;
      NumGross : UDInt;
      NumNoRead : UDInt;
      NumRead : UDInt;
      NumMatch : UDInt;
      NumMisMatch : UDInt;
   END_STRUCT;
END_TYPE

TYPE "UDT_ComMaterialReading"
VERSION : 0.1
   STRUCT
      Reading : UDInt;
      NewMaterialNumber : UDInt;
      ActualMaterialNumber : UDInt;
      NumOfTriggers : UDInt;
      NumOfReads : UDInt;
      NumOfNoReads : UDInt;
      NumOfMatches : UDInt;
      NumOfMisMatches : UDInt;
   END_STRUCT;
END_TYPE

TYPE "UDT_LatestReading"
VERSION : 0.1
   STRUCT
      ID : Int;
      Flags : Int;
      Length : Int;
      Value : Array[0..79] of Char;
   END_STRUCT;
END_TYPE

TYPE "UDT_Status"
VERSION : 0.1
   STRUCT
      EnigmaDisable : Bool;
      NoReadFault : Bool;
      MisMatchFault : Bool;
      MisTriggerFault : Bool;
      ValidData : Bool;
   END_STRUCT;
END_TYPE

TYPE "UDT_TRP_Comm"
VERSION : 0.1
   STRUCT
      NewGTIN_Number : String;
      NewBatchNumber : String;
      NewArticleNumber : UDInt;
      NewMachineID : String;
      NewBBD : String;
      ActualGTIN_Number : String;
      ActualBatchNumber : String;
      ActualAricleNumber : String;
      ActualMachineID : String;
      ActualBBD : String;
   END_STRUCT;
END_TYPE

TYPE "UDT_CON_Printer"